// TIA Portal project "FABRICA DE TAPAS - TRANSPORTE -TUNEL DE ENFRIAMIENTO" (V17) (continued)
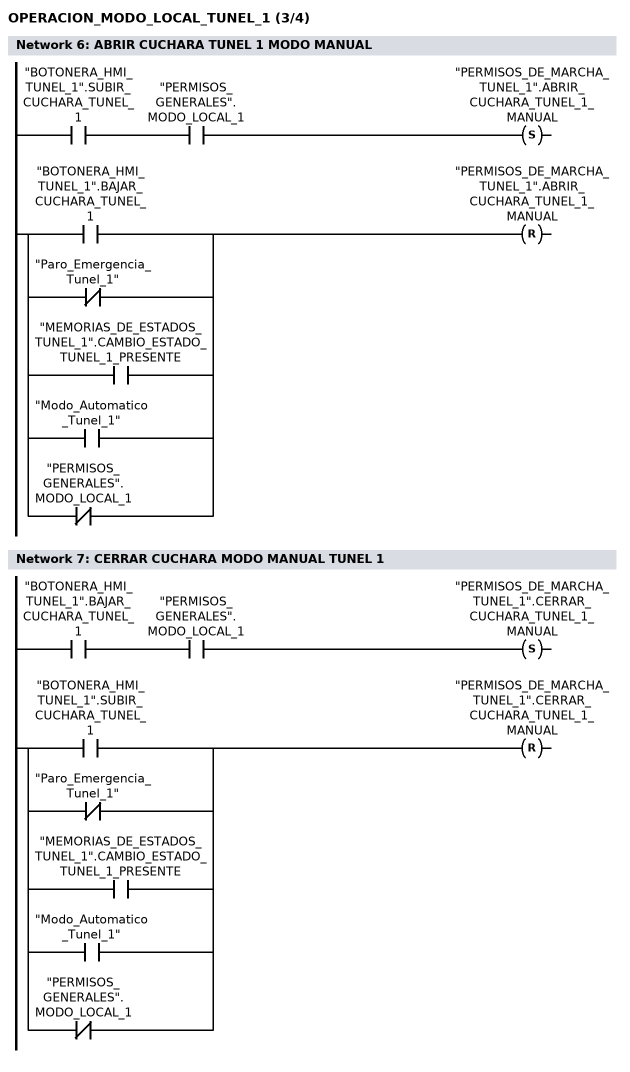
   RUNG wire#powerrail
      Contact( "BOTONERA_HMI_TUNEL_1".SUBIR_CUCHARA_TUNEL_1 )
      Contact( "PERMISOS_GENERALES".MODO_LOCAL_1 )
      S_Coil( "PERMISOS_DE_MARCHA_TUNEL_1".ABRIR_CUCHARA_TUNEL_1_MANUAL )
   END_RUNG
   RUNG wire#powerrail
      Contact( "BOTONERA_HMI_TUNEL_1".BAJAR_CUCHARA_TUNEL_1 )
      wire#w1
      R_Coil( "PERMISOS_DE_MARCHA_TUNEL_1".ABRIR_CUCHARA_TUNEL_1_MANUAL )
   END_RUNG
   RUNG wire#powerrail
      I_Contact( "Paro_Emergencia_Tunel_1" )
   END_RUNG wire#w1
   RUNG wire#powerrail
      Contact( "MEMORIAS_DE_ESTADOS_TUNEL_1".CAMBIO_ESTADO_TUNEL_1_PRESENTE )
   END_RUNG wire#w1
   RUNG wire#powerrail
      Contact( "Modo_Automatico_Tunel_1" )
   END_RUNG wire#w1
   RUNG wire#powerrail
      I_Contact( "PERMISOS_GENERALES".MODO_LOCAL_1 )
   END_RUNG wire#w1
   // the same network as SCL:
   IF "BOTONERA_HMI_TUNEL_1".SUBIR_CUCHARA_TUNEL_1 AND "PERMISOS_GENERALES".MODO_LOCAL_1 THEN
       "PERMISOS_DE_MARCHA_TUNEL_1".ABRIR_CUCHARA_TUNEL_1_MANUAL := TRUE;
   END_IF;
   IF "BOTONERA_HMI_TUNEL_1".BAJAR_CUCHARA_TUNEL_1 OR NOT "Paro_Emergencia_Tunel_1" OR "MEMORIAS_DE_ESTADOS_TUNEL_1".CAMBIO_ESTADO_TUNEL_1_PRESENTE OR "Modo_Automatico_Tunel_1" OR NOT "PERMISOS_GENERALES".MODO_LOCAL_1 THEN
       "PERMISOS_DE_MARCHA_TUNEL_1".ABRIR_CUCHARA_TUNEL_1_MANUAL := FALSE;
   END_IF;
END_REGION

REGION Network 7: CERRAR CUCHARA MODO MANUAL TUNEL 1
   RUNG wire#powerrail
      Contact( "BOTONERA_HMI_TUNEL_1".BAJAR_CUCHARA_TUNEL_1 )
      Contact( "PERMISOS_GENERALES".MODO_LOCAL_1 )
      S_Coil( "PERMISOS_DE_MARCHA_TUNEL_1".CERRAR_CUCHARA_TUNEL_1_MANUAL )
   END_RUNG
   RUNG wire#powerrail
      Contact( "BOTONERA_HMI_TUNEL_1".SUBIR_CUCHARA_TUNEL_1 )
      wire#w1
      R_Coil( "PERMISOS_DE_MARCHA_TUNEL_1".CERRAR_CUCHARA_TUNEL_1_MANUAL )
   END_RUNG
   RUNG wire#powerrail
      I_Contact( "Paro_Emergencia_Tunel_1" )
   END_RUNG wire#w1
   RUNG wire#powerrail
      Contact( "MEMORIAS_DE_ESTADOS_TUNEL_1".CAMBIO_ESTADO_TUNEL_1_PRESENTE )
   END_RUNG wire#w1
   RUNG wire#powerrail
      Contact( "Modo_Automatico_Tunel_1" )
   END_RUNG wire#w1
   RUNG wire#powerrail
      I_Contact( "PERMISOS_GENERALES".MODO_LOCAL_1 )
   END_RUNG wire#w1
   // the same network as SCL:
   IF "BOTONERA_HMI_TUNEL_1".BAJAR_CUCHARA_TUNEL_1 AND "PERMISOS_GENERALES".MODO_LOCAL_1 THEN
       "PERMISOS_DE_MARCHA_TUNEL_1".CERRAR_CUCHARA_TUNEL_1_MANUAL := TRUE;
   END_IF;
   IF "BOTONERA_HMI_TUNEL_1".SUBIR_CUCHARA_TUNEL_1 OR NOT "Paro_Emergencia_Tunel_1" OR "MEMORIAS_DE_ESTADOS_TUNEL_1".CAMBIO_ESTADO_TUNEL_1_PRESENTE OR "Modo_Automatico_Tunel_1" OR NOT "PERMISOS_GENERALES".MODO_LOCAL_1 THEN
       "PERMISOS_DE_MARCHA_TUNEL_1".CERRAR_CUCHARA_TUNEL_1_MANUAL := FALSE;
   END_IF;
END_REGION

REGION Network 8: MOVER SEPARADOR CAJAS A LA DERECHA DE MODO MANUAL TUNEL 1
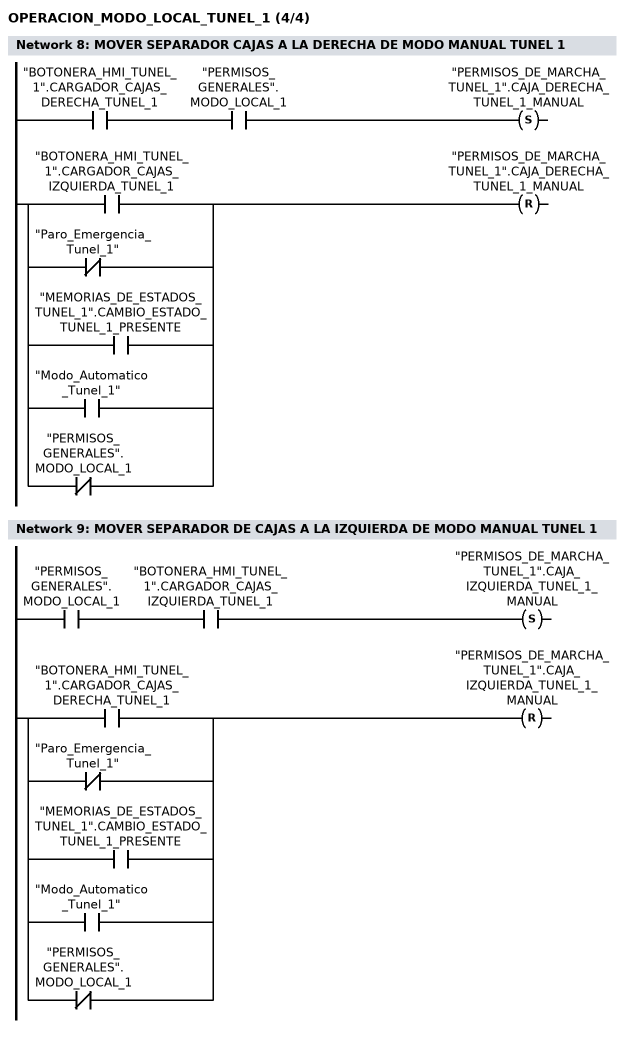
   RUNG wire#powerrail
      Contact( "BOTONERA_HMI_TUNEL_1".CARGADOR_CAJAS_DERECHA_TUNEL_1 )
      Contact( "PERMISOS_GENERALES".MODO_LOCAL_1 )
      S_Coil( "PERMISOS_DE_MARCHA_TUNEL_1".CAJA_DERECHA_TUNEL_1_MANUAL )
   END_RUNG
   RUNG wire#powerrail
      Contact( "BOTONERA_HMI_TUNEL_1".CARGADOR_CAJAS_IZQUIERDA_TUNEL_1 )
      wire#w1
      R_Coil( "PERMISOS_DE_MARCHA_TUNEL_1".CAJA_DERECHA_TUNEL_1_MANUAL )
   END_RUNG
   RUNG wire#powerrail
      I_Contact( "Paro_Emergencia_Tunel_1" )
   END_RUNG wire#w1
   RUNG wire#powerrail
      Contact( "MEMORIAS_DE_ESTADOS_TUNEL_1".CAMBIO_ESTADO_TUNEL_1_PRESENTE )
   END_RUNG wire#w1
   RUNG wire#powerrail
      Contact( "Modo_Automatico_Tunel_1" )
   END_RUNG wire#w1
   RUNG wire#powerrail
      I_Contact( "PERMISOS_GENERALES".MODO_LOCAL_1 )
   END_RUNG wire#w1
   // the same network as SCL:
   IF "BOTONERA_HMI_TUNEL_1".CARGADOR_CAJAS_DERECHA_TUNEL_1 AND "PERMISOS_GENERALES".MODO_LOCAL_1 THEN
       "PERMISOS_DE_MARCHA_TUNEL_1".CAJA_DERECHA_TUNEL_1_MANUAL := TRUE;
   END_IF;
   IF "BOTONERA_HMI_TUNEL_1".CARGADOR_CAJAS_IZQUIERDA_TUNEL_1 OR NOT "Paro_Emergencia_Tunel_1" OR "MEMORIAS_DE_ESTADOS_TUNEL_1".CAMBIO_ESTADO_TUNEL_1_PRESENTE OR "Modo_Automatico_Tunel_1" OR NOT "PERMISOS_GENERALES".MODO_LOCAL_1 THEN
       "PERMISOS_DE_MARCHA_TUNEL_1".CAJA_DERECHA_TUNEL_1_MANUAL := FALSE;
   END_IF;
END_REGION

REGION Network 9: MOVER SEPARADOR DE CAJAS A LA IZQUIERDA DE MODO MANUAL TUNEL 1
   RUNG wire#powerrail
      Contact( "PERMISOS_GENERALES".MODO_LOCAL_1 )
      Contact( "BOTONERA_HMI_TUNEL_1".CARGADOR_CAJAS_IZQUIERDA_TUNEL_1 )
      S_Coil( "PERMISOS_DE_MARCHA_TUNEL_1".CAJA_IZQUIERDA_TUNEL_1_MANUAL )
   END_RUNG
   RUNG wire#powerrail
      Contact( "BOTONERA_HMI_TUNEL_1".CARGADOR_CAJAS_DERECHA_TUNEL_1 )
      wire#w1
      R_Coil( "PERMISOS_DE_MARCHA_TUNEL_1".CAJA_IZQUIERDA_TUNEL_1_MANUAL )
   END_RUNG
   RUNG wire#powerrail
      I_Contact( "Paro_Emergencia_Tunel_1" )
   END_RUNG wire#w1
   RUNG wire#powerrail
      Contact( "MEMORIAS_DE_ESTADOS_TUNEL_1".CAMBIO_ESTADO_TUNEL_1_PRESENTE )
   END_RUNG wire#w1
   RUNG wire#powerrail
      Contact( "Modo_Automatico_Tunel_1" )
   END_RUNG wire#w1
   RUNG wire#powerrail
      I_Contact( "PERMISOS_GENERALES".MODO_LOCAL_1 )
   END_RUNG wire#w1
   // the same network as SCL:
   IF "PERMISOS_GENERALES".MODO_LOCAL_1 AND "BOTONERA_HMI_TUNEL_1".CARGADOR_CAJAS_IZQUIERDA_TUNEL_1 THEN
       "PERMISOS_DE_MARCHA_TUNEL_1".CAJA_IZQUIERDA_TUNEL_1_MANUAL := TRUE;
   END_IF;
   IF "BOTONERA_HMI_TUNEL_1".CARGADOR_CAJAS_DERECHA_TUNEL_1 OR NOT "Paro_Emergencia_Tunel_1" OR "MEMORIAS_DE_ESTADOS_TUNEL_1".CAMBIO_ESTADO_TUNEL_1_PRESENTE OR "Modo_Automatico_Tunel_1" OR NOT "PERMISOS_GENERALES".MODO_LOCAL_1 THEN
       "PERMISOS_DE_MARCHA_TUNEL_1".CAJA_IZQUIERDA_TUNEL_1_MANUAL := FALSE;
   END_IF;
END_REGION
END_FUNCTION

FUNCTION "OPERACION_MODO_LOCAL_TUNEL_2" : Void   // FC4, LAD
{ S7_Optimized_Access := 'TRUE' }
VERSION : 0.1
BEGIN

REGION Network 1
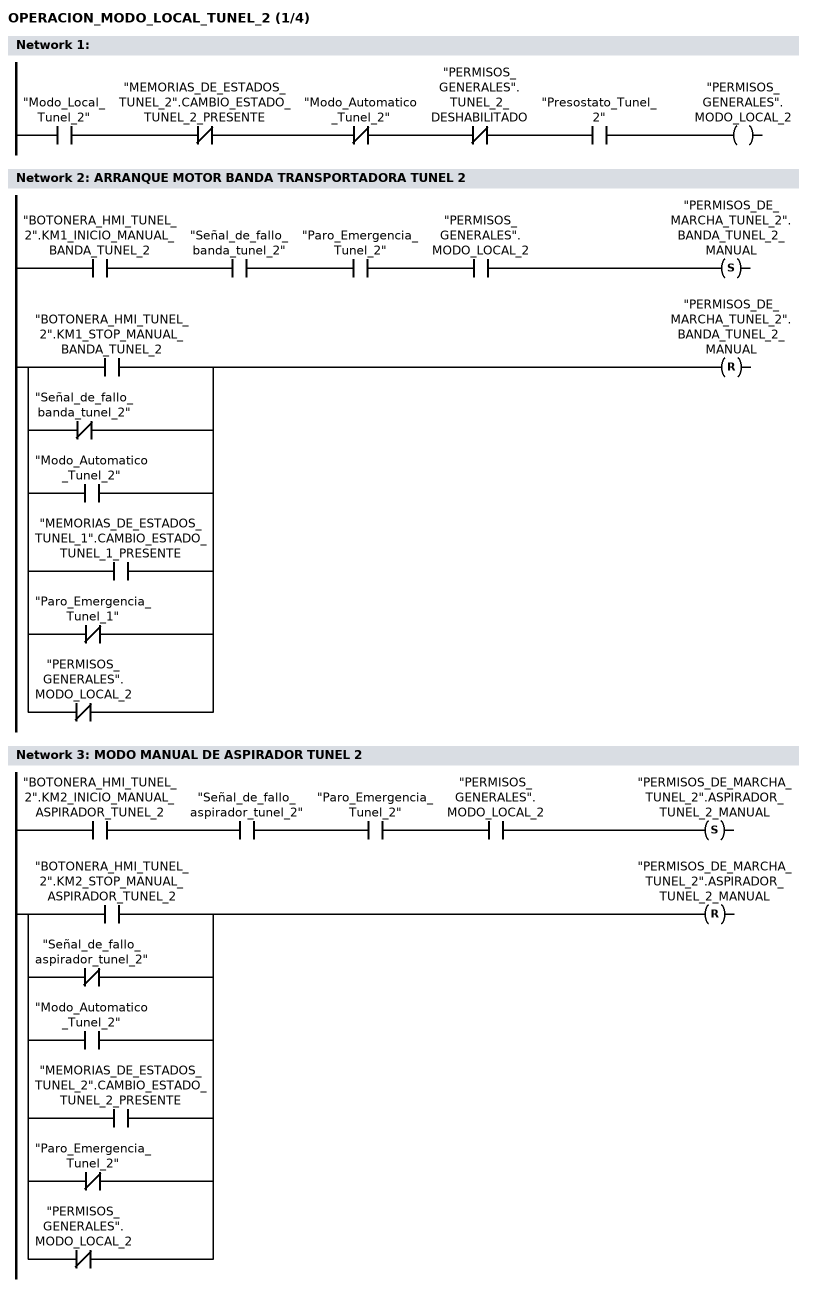
   RUNG wire#powerrail
      Contact( "Modo_Local_Tunel_2" )
      I_Contact( "MEMORIAS_DE_ESTADOS_TUNEL_2".CAMBIO_ESTADO_TUNEL_2_PRESENTE )
      I_Contact( "Modo_Automatico_Tunel_2" )
      I_Contact( "PERMISOS_GENERALES".TUNEL_2_DESHABILITADO )
      Contact( "Presostato_Tunel_2" )
      Coil( "PERMISOS_GENERALES".MODO_LOCAL_2 )
   END_RUNG
   // the same network as SCL:
   "PERMISOS_GENERALES".MODO_LOCAL_2 := "Modo_Local_Tunel_2" AND NOT "MEMORIAS_DE_ESTADOS_TUNEL_2".CAMBIO_ESTADO_TUNEL_2_PRESENTE AND NOT "Modo_Automatico_Tunel_2" AND NOT "PERMISOS_GENERALES".TUNEL_2_DESHABILITADO AND "Presostato_Tunel_2";
END_REGION

REGION Network 2: ARRANQUE MOTOR BANDA TRANSPORTADORA TUNEL 2
   RUNG wire#powerrail
      Contact( "BOTONERA_HMI_TUNEL_2".KM1_INICIO_MANUAL_BANDA_TUNEL_2 )
      Contact( "Señal_de_fallo_banda_tunel_2" )
      Contact( "Paro_Emergencia_Tunel_2" )
      Contact( "PERMISOS_GENERALES".MODO_LOCAL_2 )
      S_Coil( "PERMISOS_DE_MARCHA_TUNEL_2".BANDA_TUNEL_2_MANUAL )
   END_RUNG
   RUNG wire#powerrail
      Contact( "BOTONERA_HMI_TUNEL_2".KM1_STOP_MANUAL_BANDA_TUNEL_2 )
      wire#w1
      R_Coil( "PERMISOS_DE_MARCHA_TUNEL_2".BANDA_TUNEL_2_MANUAL )
   END_RUNG
   RUNG wire#powerrail
      I_Contact( "Señal_de_fallo_banda_tunel_2" )
   END_RUNG wire#w1
   RUNG wire#powerrail
      Contact( "Modo_Automatico_Tunel_2" )
   END_RUNG wire#w1
   RUNG wire#powerrail
      Contact( "MEMORIAS_DE_ESTADOS_TUNEL_1".CAMBIO_ESTADO_TUNEL_1_PRESENTE )
   END_RUNG wire#w1
   RUNG wire#powerrail
      I_Contact( "Paro_Emergencia_Tunel_1" )
   END_RUNG wire#w1
   RUNG wire#powerrail
      I_Contact( "PERMISOS_GENERALES".MODO_LOCAL_2 )
   END_RUNG wire#w1
   // the same network as SCL:
   IF "BOTONERA_HMI_TUNEL_2".KM1_INICIO_MANUAL_BANDA_TUNEL_2 AND "Señal_de_fallo_banda_tunel_2" AND "Paro_Emergencia_Tunel_2" AND "PERMISOS_GENERALES".MODO_LOCAL_2 THEN
       "PERMISOS_DE_MARCHA_TUNEL_2".BANDA_TUNEL_2_MANUAL := TRUE;
   END_IF;
   IF "BOTONERA_HMI_TUNEL_2".KM1_STOP_MANUAL_BANDA_TUNEL_2 OR NOT "Señal_de_fallo_banda_tunel_2" OR "Modo_Automatico_Tunel_2" OR "MEMORIAS_DE_ESTADOS_TUNEL_1".CAMBIO_ESTADO_TUNEL_1_PRESENTE OR NOT "Paro_Emergencia_Tunel_1" OR NOT "PERMISOS_GENERALES".MODO_LOCAL_2 THEN
       "PERMISOS_DE_MARCHA_TUNEL_2".BANDA_TUNEL_2_MANUAL := FALSE;
   END_IF;
END_REGION

REGION Network 3: MODO MANUAL DE ASPIRADOR TUNEL 2
   RUNG wire#powerrail
      Contact( "BOTONERA_HMI_TUNEL_2".KM2_INICIO_MANUAL_ASPIRADOR_TUNEL_2 )
      Contact( "Señal_de_fallo_aspirador_tunel_2" )
      Contact( "Paro_Emergencia_Tunel_2" )
      Contact( "PERMISOS_GENERALES".MODO_LOCAL_2 )
      S_Coil( "PERMISOS_DE_MARCHA_TUNEL_2".ASPIRADOR_TUNEL_2_MANUAL )
   END_RUNG
   RUNG wire#powerrail
      Contact( "BOTONERA_HMI_TUNEL_2".KM2_STOP_MANUAL_ASPIRADOR_TUNEL_2 )
      wire#w1
      R_Coil( "PERMISOS_DE_MARCHA_TUNEL_2".ASPIRADOR_TUNEL_2_MANUAL )
   END_RUNG
   RUNG wire#powerrail
      I_Contact( "Señal_de_fallo_aspirador_tunel_2" )
   END_RUNG wire#w1
   RUNG wire#powerrail
      Contact( "Modo_Automatico_Tunel_2" )
   END_RUNG wire#w1
   RUNG wire#powerrail
      Contact( "MEMORIAS_DE_ESTADOS_TUNEL_2".CAMBIO_ESTADO_TUNEL_2_PRESENTE )
   END_RUNG wire#w1
   RUNG wire#powerrail
      I_Contact( "Paro_Emergencia_Tunel_2" )
   END_RUNG wire#w1
   RUNG wire#powerrail
      I_Contact( "PERMISOS_GENERALES".MODO_LOCAL_2 )
   END_RUNG wire#w1
   // the same network as SCL:
   IF "BOTONERA_HMI_TUNEL_2".KM2_INICIO_MANUAL_ASPIRADOR_TUNEL_2 AND "Señal_de_fallo_aspirador_tunel_2" AND "Paro_Emergencia_Tunel_2" AND "PERMISOS_GENERALES".MODO_LOCAL_2 THEN
       "PERMISOS_DE_MARCHA_TUNEL_2".ASPIRADOR_TUNEL_2_MANUAL := TRUE;
   END_IF;
   IF "BOTONERA_HMI_TUNEL_2".KM2_STOP_MANUAL_ASPIRADOR_TUNEL_2 OR NOT "Señal_de_fallo_aspirador_tunel_2" OR "Modo_Automatico_Tunel_2" OR "MEMORIAS_DE_ESTADOS_TUNEL_2".CAMBIO_ESTADO_TUNEL_2_PRESENTE OR NOT "Paro_Emergencia_Tunel_2" OR NOT "PERMISOS_GENERALES".MODO_LOCAL_2 THEN
       "PERMISOS_DE_MARCHA_TUNEL_2".ASPIRADOR_TUNEL_2_MANUAL := FALSE;
   END_IF;
END_REGION

REGION Network 4: MODO MANUAL VENTILADOR TUNEL 2
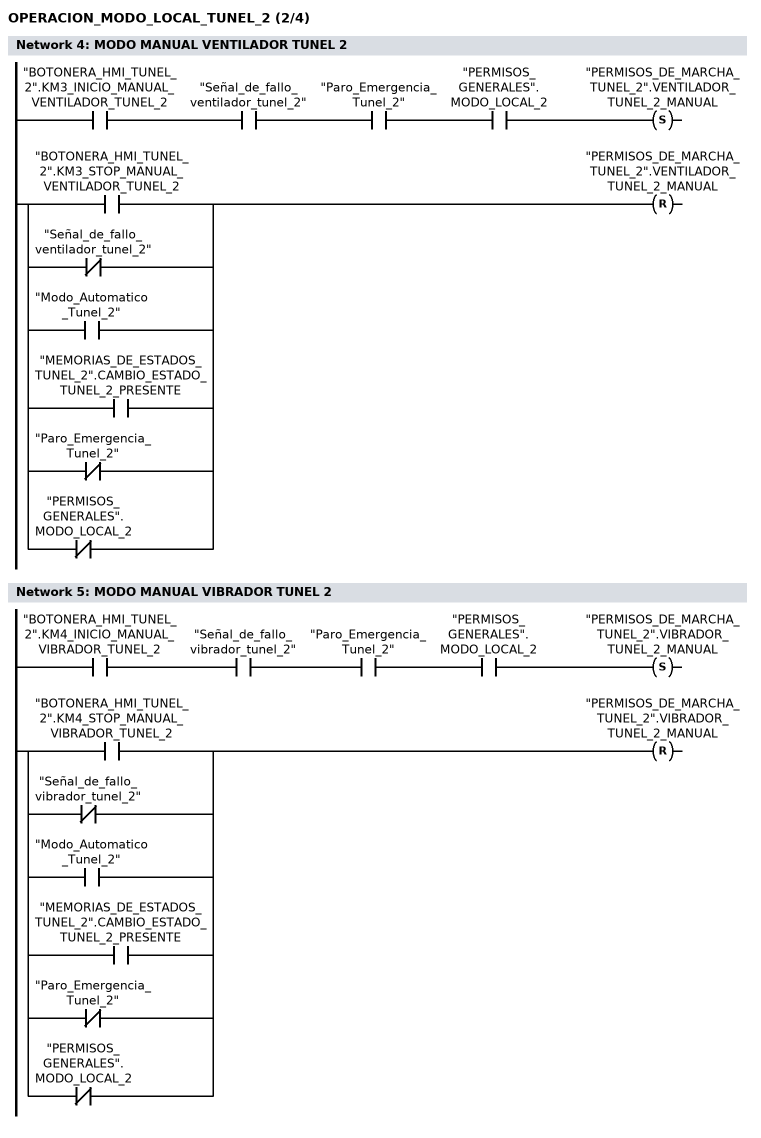
   RUNG wire#powerrail
      Contact( "BOTONERA_HMI_TUNEL_2".KM3_INICIO_MANUAL_VENTILADOR_TUNEL_2 )
      Contact( "Señal_de_fallo_ventilador_tunel_2" )
      Contact( "Paro_Emergencia_Tunel_2" )
      Contact( "PERMISOS_GENERALES".MODO_LOCAL_2 )
      S_Coil( "PERMISOS_DE_MARCHA_TUNEL_2".VENTILADOR_TUNEL_2_MANUAL )
   END_RUNG
   RUNG wire#powerrail
      Contact( "BOTONERA_HMI_TUNEL_2".KM3_STOP_MANUAL_VENTILADOR_TUNEL_2 )
      wire#w1
      R_Coil( "PERMISOS_DE_MARCHA_TUNEL_2".VENTILADOR_TUNEL_2_MANUAL )
   END_RUNG
   RUNG wire#powerrail
      I_Contact( "Señal_de_fallo_ventilador_tunel_2" )
   END_RUNG wire#w1
   RUNG wire#powerrail
      Contact( "Modo_Automatico_Tunel_2" )
   END_RUNG wire#w1
   RUNG wire#powerrail
      Contact( "MEMORIAS_DE_ESTADOS_TUNEL_2".CAMBIO_ESTADO_TUNEL_2_PRESENTE )
   END_RUNG wire#w1
   RUNG wire#powerrail
      I_Contact( "Paro_Emergencia_Tunel_2" )
   END_RUNG wire#w1
   RUNG wire#powerrail
      I_Contact( "PERMISOS_GENERALES".MODO_LOCAL_2 )
   END_RUNG wire#w1
   // the same network as SCL:
   IF "BOTONERA_HMI_TUNEL_2".KM3_INICIO_MANUAL_VENTILADOR_TUNEL_2 AND "Señal_de_fallo_ventilador_tunel_2" AND "Paro_Emergencia_Tunel_2" AND "PERMISOS_GENERALES".MODO_LOCAL_2 THEN
       "PERMISOS_DE_MARCHA_TUNEL_2".VENTILADOR_TUNEL_2_MANUAL := TRUE;
   END_IF;
   IF "BOTONERA_HMI_TUNEL_2".KM3_STOP_MANUAL_VENTILADOR_TUNEL_2 OR NOT "Señal_de_fallo_ventilador_tunel_2" OR "Modo_Automatico_Tunel_2" OR "MEMORIAS_DE_ESTADOS_TUNEL_2".CAMBIO_ESTADO_TUNEL_2_PRESENTE OR NOT "Paro_Emergencia_Tunel_2" OR NOT "PERMISOS_GENERALES".MODO_LOCAL_2 THEN
       "PERMISOS_DE_MARCHA_TUNEL_2".VENTILADOR_TUNEL_2_MANUAL := FALSE;
   END_IF;
END_REGION

REGION Network 5: MODO MANUAL VIBRADOR TUNEL 2
   RUNG wire#powerrail
      Contact( "BOTONERA_HMI_TUNEL_2".KM4_INICIO_MANUAL_VIBRADOR_TUNEL_2 )
      Contact( "Señal_de_fallo_vibrador_tunel_2" )
      Contact( "Paro_Emergencia_Tunel_2" )
      Contact( "PERMISOS_GENERALES".MODO_LOCAL_2 )
      S_Coil( "PERMISOS_DE_MARCHA_TUNEL_2".VIBRADOR_TUNEL_2_MANUAL )
   END_RUNG
   RUNG wire#powerrail
      Contact( "BOTONERA_HMI_TUNEL_2".KM4_STOP_MANUAL_VIBRADOR_TUNEL_2 )
      wire#w1
      R_Coil( "PERMISOS_DE_MARCHA_TUNEL_2".VIBRADOR_TUNEL_2_MANUAL )
   END_RUNG
   RUNG wire#powerrail
      I_Contact( "Señal_de_fallo_vibrador_tunel_2" )
   END_RUNG wire#w1
   RUNG wire#powerrail
      Contact( "Modo_Automatico_Tunel_2" )
   END_RUNG wire#w1
   RUNG wire#powerrail
      Contact( "MEMORIAS_DE_ESTADOS_TUNEL_2".CAMBIO_ESTADO_TUNEL_2_PRESENTE )
   END_RUNG wire#w1
   RUNG wire#powerrail
      I_Contact( "Paro_Emergencia_Tunel_2" )
   END_RUNG wire#w1
   RUNG wire#powerrail
      I_Contact( "PERMISOS_GENERALES".MODO_LOCAL_2 )
   END_RUNG wire#w1
   // the same network as SCL:
   IF "BOTONERA_HMI_TUNEL_2".KM4_INICIO_MANUAL_VIBRADOR_TUNEL_2 AND "Señal_de_fallo_vibrador_tunel_2" AND "Paro_Emergencia_Tunel_2" AND "PERMISOS_GENERALES".MODO_LOCAL_2 THEN
       "PERMISOS_DE_MARCHA_TUNEL_2".VIBRADOR_TUNEL_2_MANUAL := TRUE;
   END_IF;
   IF "BOTONERA_HMI_TUNEL_2".KM4_STOP_MANUAL_VIBRADOR_TUNEL_2 OR NOT "Señal_de_fallo_vibrador_tunel_2" OR "Modo_Automatico_Tunel_2" OR "MEMORIAS_DE_ESTADOS_TUNEL_2".CAMBIO_ESTADO_TUNEL_2_PRESENTE OR NOT "Paro_Emergencia_Tunel_2" OR NOT "PERMISOS_GENERALES".MODO_LOCAL_2 THEN
       "PERMISOS_DE_MARCHA_TUNEL_2".VIBRADOR_TUNEL_2_MANUAL := FALSE;
   END_IF;
END_REGION

REGION Network 6: ABRIR CUCHARA TUNEL 2 MODO MANUAL
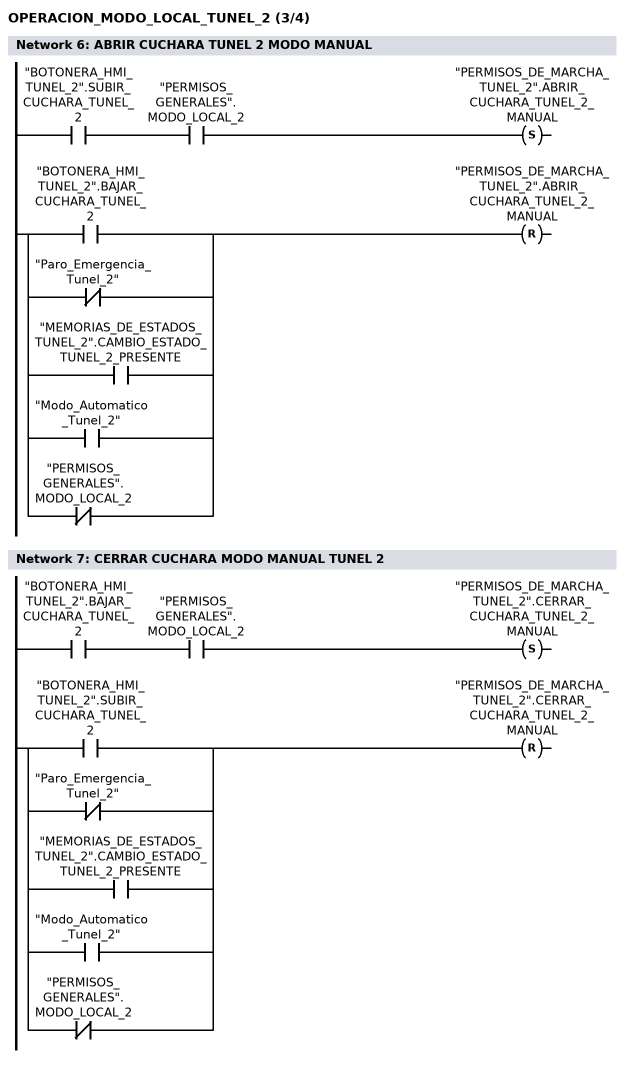
   RUNG wire#powerrail
      Contact( "BOTONERA_HMI_TUNEL_2".SUBIR_CUCHARA_TUNEL_2 )
      Contact( "PERMISOS_GENERALES".MODO_LOCAL_2 )
      S_Coil( "PERMISOS_DE_MARCHA_TUNEL_2".ABRIR_CUCHARA_TUNEL_2_MANUAL )
   END_RUNG
   RUNG wire#powerrail
      Contact( "BOTONERA_HMI_TUNEL_2".BAJAR_CUCHARA_TUNEL_2 )
      wire#w1
      R_Coil( "PERMISOS_DE_MARCHA_TUNEL_2".ABRIR_CUCHARA_TUNEL_2_MANUAL )
   END_RUNG
   RUNG wire#powerrail
      I_Contact( "Paro_Emergencia_Tunel_2" )
   END_RUNG wire#w1
   RUNG wire#powerrail
      Contact( "MEMORIAS_DE_ESTADOS_TUNEL_2".CAMBIO_ESTADO_TUNEL_2_PRESENTE )
   END_RUNG wire#w1
   RUNG wire#powerrail
      Contact( "Modo_Automatico_Tunel_2" )
   END_RUNG wire#w1
   RUNG wire#powerrail
      I_Contact( "PERMISOS_GENERALES".MODO_LOCAL_2 )
   END_RUNG wire#w1
   // the same network as SCL:
   IF "BOTONERA_HMI_TUNEL_2".SUBIR_CUCHARA_TUNEL_2 AND "PERMISOS_GENERALES".MODO_LOCAL_2 THEN
       "PERMISOS_DE_MARCHA_TUNEL_2".ABRIR_CUCHARA_TUNEL_2_MANUAL := TRUE;
   END_IF;
   IF "BOTONERA_HMI_TUNEL_2".BAJAR_CUCHARA_TUNEL_2 OR NOT "Paro_Emergencia_Tunel_2" OR "MEMORIAS_DE_ESTADOS_TUNEL_2".CAMBIO_ESTADO_TUNEL_2_PRESENTE OR "Modo_Automatico_Tunel_2" OR NOT "PERMISOS_GENERALES".MODO_LOCAL_2 THEN
       "PERMISOS_DE_MARCHA_TUNEL_2".ABRIR_CUCHARA_TUNEL_2_MANUAL := FALSE;
   END_IF;
END_REGION

REGION Network 7: CERRAR CUCHARA MODO MANUAL TUNEL 2
   RUNG wire#powerrail
      Contact( "BOTONERA_HMI_TUNEL_2".BAJAR_CUCHARA_TUNEL_2 )
      Contact( "PERMISOS_GENERALES".MODO_LOCAL_2 )
      S_Coil( "PERMISOS_DE_MARCHA_TUNEL_2".CERRAR_CUCHARA_TUNEL_2_MANUAL )
   END_RUNG
   RUNG wire#powerrail
      Contact( "BOTONERA_HMI_TUNEL_2".SUBIR_CUCHARA_TUNEL_2 )
      wire#w1
      R_Coil( "PERMISOS_DE_MARCHA_TUNEL_2".CERRAR_CUCHARA_TUNEL_2_MANUAL )
   END_RUNG
   RUNG wire#powerrail
      I_Contact( "Paro_Emergencia_Tunel_2" )
   END_RUNG wire#w1
   RUNG wire#powerrail
      Contact( "MEMORIAS_DE_ESTADOS_TUNEL_2".CAMBIO_ESTADO_TUNEL_2_PRESENTE )
   END_RUNG wire#w1
   RUNG wire#powerrail
      Contact( "Modo_Automatico_Tunel_2" )
   END_RUNG wire#w1
   RUNG wire#powerrail
      I_Contact( "PERMISOS_GENERALES".MODO_LOCAL_2 )
   END_RUNG wire#w1
   // the same network as SCL:
   IF "BOTONERA_HMI_TUNEL_2".BAJAR_CUCHARA_TUNEL_2 AND "PERMISOS_GENERALES".MODO_LOCAL_2 THEN
       "PERMISOS_DE_MARCHA_TUNEL_2".CERRAR_CUCHARA_TUNEL_2_MANUAL := TRUE;
   END_IF;
   IF "BOTONERA_HMI_TUNEL_2".SUBIR_CUCHARA_TUNEL_2 OR NOT "Paro_Emergencia_Tunel_2" OR "MEMORIAS_DE_ESTADOS_TUNEL_2".CAMBIO_ESTADO_TUNEL_2_PRESENTE OR "Modo_Automatico_Tunel_2" OR NOT "PERMISOS_GENERALES".MODO_LOCAL_2 THEN
       "PERMISOS_DE_MARCHA_TUNEL_2".CERRAR_CUCHARA_TUNEL_2_MANUAL := FALSE;
   END_IF;
END_REGION

REGION Network 8: MOVER SEPARADOR CAJAS A LA DERECHA DE MODO MANUAL TUNEL 2
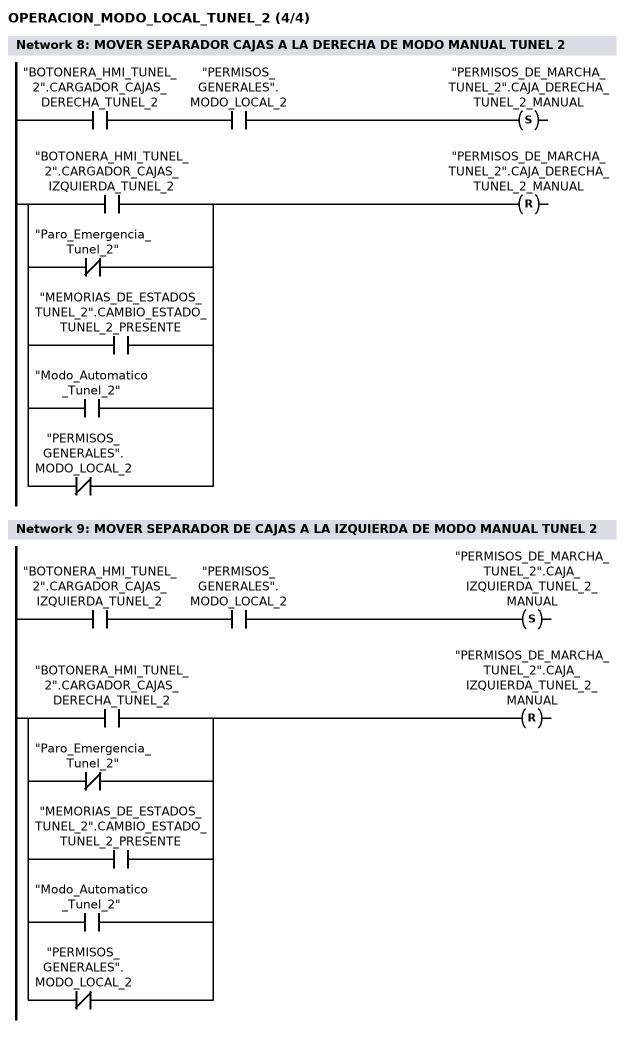
   RUNG wire#powerrail
      Contact( "BOTONERA_HMI_TUNEL_2".CARGADOR_CAJAS_DERECHA_TUNEL_2 )
      Contact( "PERMISOS_GENERALES".MODO_LOCAL_2 )
      S_Coil( "PERMISOS_DE_MARCHA_TUNEL_2".CAJA_DERECHA_TUNEL_2_MANUAL )
   END_RUNG
   RUNG wire#powerrail
      Contact( "BOTONERA_HMI_TUNEL_2".CARGADOR_CAJAS_IZQUIERDA_TUNEL_2 )
      wire#w1
      R_Coil( "PERMISOS_DE_MARCHA_TUNEL_2".CAJA_DERECHA_TUNEL_2_MANUAL )
   END_RUNG
   RUNG wire#powerrail
      I_Contact( "Paro_Emergencia_Tunel_2" )
   END_RUNG wire#w1
   RUNG wire#powerrail
      Contact( "MEMORIAS_DE_ESTADOS_TUNEL_2".CAMBIO_ESTADO_TUNEL_2_PRESENTE )
   END_RUNG wire#w1
   RUNG wire#powerrail
      Contact( "Modo_Automatico_Tunel_2" )
   END_RUNG wire#w1
   RUNG wire#powerrail
      I_Contact( "PERMISOS_GENERALES".MODO_LOCAL_2 )
   END_RUNG wire#w1
   // the same network as SCL:
   IF "BOTONERA_HMI_TUNEL_2".CARGADOR_CAJAS_DERECHA_TUNEL_2 AND "PERMISOS_GENERALES".MODO_LOCAL_2 THEN
       "PERMISOS_DE_MARCHA_TUNEL_2".CAJA_DERECHA_TUNEL_2_MANUAL := TRUE;
   END_IF;
   IF "BOTONERA_HMI_TUNEL_2".CARGADOR_CAJAS_IZQUIERDA_TUNEL_2 OR NOT "Paro_Emergencia_Tunel_2" OR "MEMORIAS_DE_ESTADOS_TUNEL_2".CAMBIO_ESTADO_TUNEL_2_PRESENTE OR "Modo_Automatico_Tunel_2" OR NOT "PERMISOS_GENERALES".MODO_LOCAL_2 THEN
       "PERMISOS_DE_MARCHA_TUNEL_2".CAJA_DERECHA_TUNEL_2_MANUAL := FALSE;
   END_IF;
END_REGION

REGION Network 9: MOVER SEPARADOR DE CAJAS A LA IZQUIERDA DE MODO MANUAL TUNEL 2
   RUNG wire#powerrail
      Contact( "BOTONERA_HMI_TUNEL_2".CARGADOR_CAJAS_IZQUIERDA_TUNEL_2 )
      Contact( "PERMISOS_GENERALES".MODO_LOCAL_2 )
      S_Coil( "PERMISOS_DE_MARCHA_TUNEL_2".CAJA_IZQUIERDA_TUNEL_2_MANUAL )
   END_RUNG
   RUNG wire#powerrail
      Contact( "BOTONERA_HMI_TUNEL_2".CARGADOR_CAJAS_DERECHA_TUNEL_2 )
      wire#w1
      R_Coil( "PERMISOS_DE_MARCHA_TUNEL_2".CAJA_IZQUIERDA_TUNEL_2_MANUAL )
   END_RUNG
   RUNG wire#powerrail
      I_Contact( "Paro_Emergencia_Tunel_2" )
   END_RUNG wire#w1
   RUNG wire#powerrail
      Contact( "MEMORIAS_DE_ESTADOS_TUNEL_2".CAMBIO_ESTADO_TUNEL_2_PRESENTE )
   END_RUNG wire#w1
   RUNG wire#powerrail
      Contact( "Modo_Automatico_Tunel_2" )
   END_RUNG wire#w1
   RUNG wire#powerrail
      I_Contact( "PERMISOS_GENERALES".MODO_LOCAL_2 )
   END_RUNG wire#w1
   // the same network as SCL:
   IF "BOTONERA_HMI_TUNEL_2".CARGADOR_CAJAS_IZQUIERDA_TUNEL_2 AND "PERMISOS_GENERALES".MODO_LOCAL_2 THEN
       "PERMISOS_DE_MARCHA_TUNEL_2".CAJA_IZQUIERDA_TUNEL_2_MANUAL := TRUE;
   END_IF;
   IF "BOTONERA_HMI_TUNEL_2".CARGADOR_CAJAS_DERECHA_TUNEL_2 OR NOT "Paro_Emergencia_Tunel_2" OR "MEMORIAS_DE_ESTADOS_TUNEL_2".CAMBIO_ESTADO_TUNEL_2_PRESENTE OR "Modo_Automatico_Tunel_2" OR NOT "PERMISOS_GENERALES".MODO_LOCAL_2 THEN
       "PERMISOS_DE_MARCHA_TUNEL_2".CAJA_IZQUIERDA_TUNEL_2_MANUAL := FALSE;
   END_IF;
END_REGION
END_FUNCTION

FUNCTION "OPERACION_MANUAL_TRANSPORTE" : Void   // FC5, LAD
{ S7_Optimized_Access := 'TRUE' }
VERSION : 0.1
BEGIN

REGION Network 1
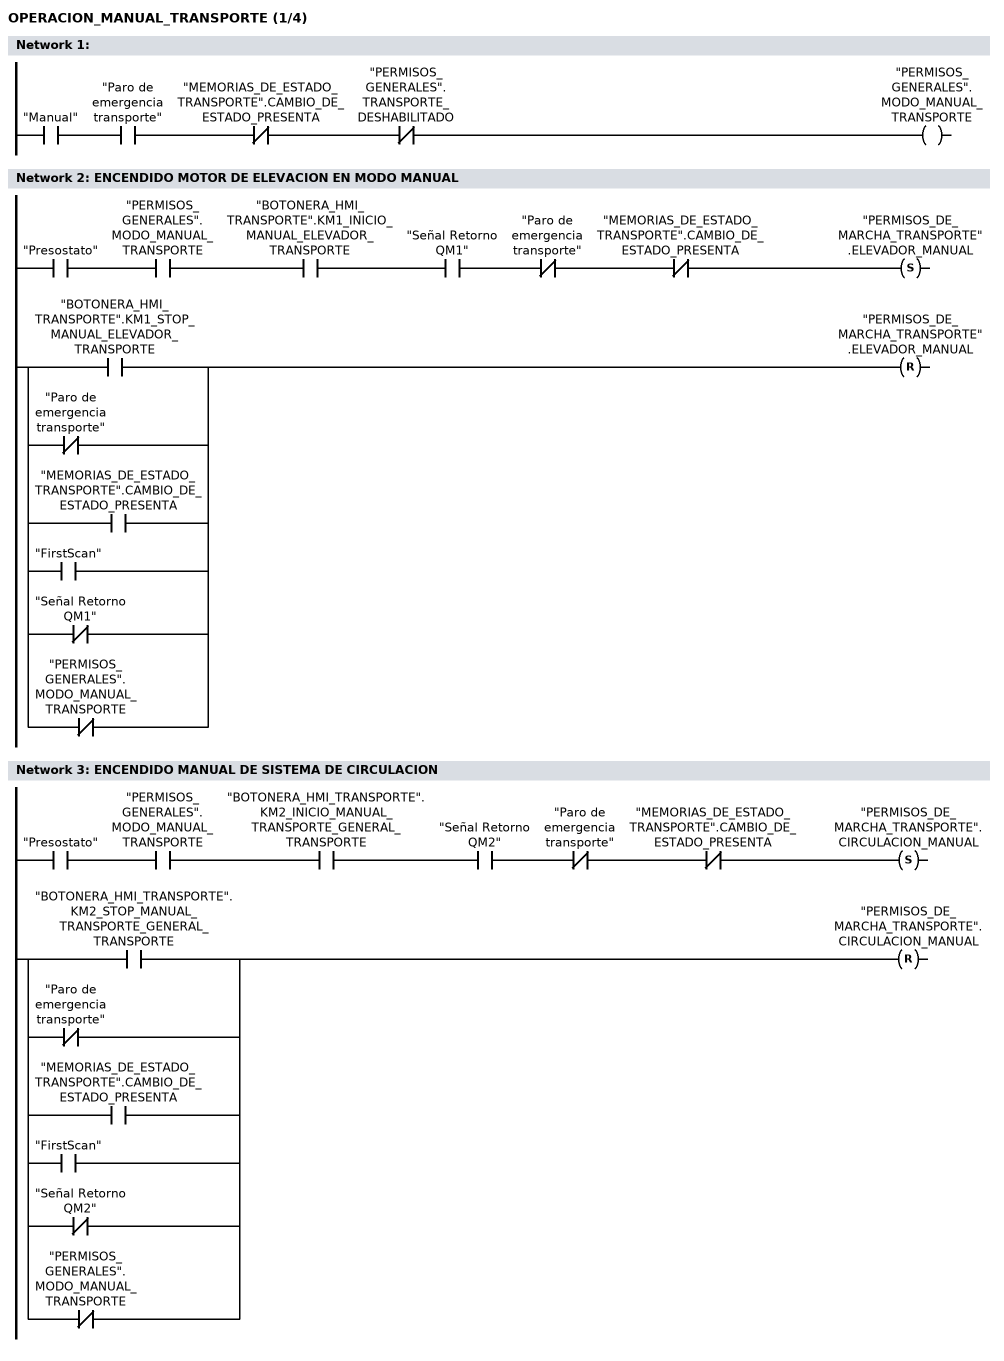
   RUNG wire#powerrail
      Contact( "Manual" )
      Contact( "Paro de emergencia transporte" )
      I_Contact( "MEMORIAS_DE_ESTADO_TRANSPORTE".CAMBIO_DE_ESTADO_PRESENTA )
      I_Contact( "PERMISOS_GENERALES".TRANSPORTE_DESHABILITADO )
      Coil( "PERMISOS_GENERALES".MODO_MANUAL_TRANSPORTE )
   END_RUNG
   // the same network as SCL:
   "PERMISOS_GENERALES".MODO_MANUAL_TRANSPORTE := "Manual" AND "Paro de emergencia transporte" AND NOT "MEMORIAS_DE_ESTADO_TRANSPORTE".CAMBIO_DE_ESTADO_PRESENTA AND NOT "PERMISOS_GENERALES".TRANSPORTE_DESHABILITADO;
END_REGION

REGION Network 2: ENCENDIDO MOTOR DE ELEVACION EN MODO MANUAL
   RUNG wire#powerrail
      Contact( "Presostato" )
      Contact( "PERMISOS_GENERALES".MODO_MANUAL_TRANSPORTE )
      Contact( "BOTONERA_HMI_TRANSPORTE".KM1_INICIO_MANUAL_ELEVADOR_TRANSPORTE )
      Contact( "Señal Retorno QM1" )
      I_Contact( "Paro de emergencia transporte" )
      I_Contact( "MEMORIAS_DE_ESTADO_TRANSPORTE".CAMBIO_DE_ESTADO_PRESENTA )
      S_Coil( "PERMISOS_DE_MARCHA_TRANSPORTE".ELEVADOR_MANUAL )
   END_RUNG
   RUNG wire#powerrail
      Contact( "BOTONERA_HMI_TRANSPORTE".KM1_STOP_MANUAL_ELEVADOR_TRANSPORTE )
      wire#w1
      R_Coil( "PERMISOS_DE_MARCHA_TRANSPORTE".ELEVADOR_MANUAL )
   END_RUNG
   RUNG wire#powerrail
      I_Contact( "Paro de emergencia transporte" )
   END_RUNG wire#w1
   RUNG wire#powerrail
      Contact( "MEMORIAS_DE_ESTADO_TRANSPORTE".CAMBIO_DE_ESTADO_PRESENTA )
   END_RUNG wire#w1
   RUNG wire#powerrail
      Contact( "FirstScan" )
   END_RUNG wire#w1
   RUNG wire#powerrail
      I_Contact( "Señal Retorno QM1" )
   END_RUNG wire#w1
   RUNG wire#powerrail
      I_Contact( "PERMISOS_GENERALES".MODO_MANUAL_TRANSPORTE )
   END_RUNG wire#w1
   // the same network as SCL:
   IF "Presostato" AND "PERMISOS_GENERALES".MODO_MANUAL_TRANSPORTE AND "BOTONERA_HMI_TRANSPORTE".KM1_INICIO_MANUAL_ELEVADOR_TRANSPORTE AND "Señal Retorno QM1" AND NOT "Paro de emergencia transporte" AND NOT "MEMORIAS_DE_ESTADO_TRANSPORTE".CAMBIO_DE_ESTADO_PRESENTA THEN
       "PERMISOS_DE_MARCHA_TRANSPORTE".ELEVADOR_MANUAL := TRUE;
   END_IF;
   IF "BOTONERA_HMI_TRANSPORTE".KM1_STOP_MANUAL_ELEVADOR_TRANSPORTE OR NOT "Paro de emergencia transporte" OR "MEMORIAS_DE_ESTADO_TRANSPORTE".CAMBIO_DE_ESTADO_PRESENTA OR "FirstScan" OR NOT "Señal Retorno QM1" OR NOT "PERMISOS_GENERALES".MODO_MANUAL_TRANSPORTE THEN
       "PERMISOS_DE_MARCHA_TRANSPORTE".ELEVADOR_MANUAL := FALSE;
   END_IF;
END_REGION

REGION Network 3: ENCENDIDO MANUAL DE SISTEMA DE CIRCULACION
   RUNG wire#powerrail
      Contact( "Presostato" )
      Contact( "PERMISOS_GENERALES".MODO_MANUAL_TRANSPORTE )
      Contact( "BOTONERA_HMI_TRANSPORTE".KM2_INICIO_MANUAL_TRANSPORTE_GENERAL_TRANSPORTE )
      Contact( "Señal Retorno QM2" )
      I_Contact( "Paro de emergencia transporte" )
      I_Contact( "MEMORIAS_DE_ESTADO_TRANSPORTE".CAMBIO_DE_ESTADO_PRESENTA )
      S_Coil( "PERMISOS_DE_MARCHA_TRANSPORTE".CIRCULACION_MANUAL )
   END_RUNG
   RUNG wire#powerrail
      Contact( "BOTONERA_HMI_TRANSPORTE".KM2_STOP_MANUAL_TRANSPORTE_GENERAL_TRANSPORTE )
      wire#w1
      R_Coil( "PERMISOS_DE_MARCHA_TRANSPORTE".CIRCULACION_MANUAL )
   END_RUNG
   RUNG wire#powerrail
      I_Contact( "Paro de emergencia transporte" )
   END_RUNG wire#w1
   RUNG wire#powerrail
      Contact( "MEMORIAS_DE_ESTADO_TRANSPORTE".CAMBIO_DE_ESTADO_PRESENTA )
   END_RUNG wire#w1
   RUNG wire#powerrail
      Contact( "FirstScan" )
   END_RUNG wire#w1
   RUNG wire#powerrail
      I_Contact( "Señal Retorno QM2" )
   END_RUNG wire#w1
   RUNG wire#powerrail
      I_Contact( "PERMISOS_GENERALES".MODO_MANUAL_TRANSPORTE )
   END_RUNG wire#w1
   // the same network as SCL:
   IF "Presostato" AND "PERMISOS_GENERALES".MODO_MANUAL_TRANSPORTE AND "BOTONERA_HMI_TRANSPORTE".KM2_INICIO_MANUAL_TRANSPORTE_GENERAL_TRANSPORTE AND "Señal Retorno QM2" AND NOT "Paro de emergencia transporte" AND NOT "MEMORIAS_DE_ESTADO_TRANSPORTE".CAMBIO_DE_ESTADO_PRESENTA THEN
       "PERMISOS_DE_MARCHA_TRANSPORTE".CIRCULACION_MANUAL := TRUE;
   END_IF;
   IF "BOTONERA_HMI_TRANSPORTE".KM2_STOP_MANUAL_TRANSPORTE_GENERAL_TRANSPORTE OR NOT "Paro de emergencia transporte" OR "MEMORIAS_DE_ESTADO_TRANSPORTE".CAMBIO_DE_ESTADO_PRESENTA OR "FirstScan" OR NOT "Señal Retorno QM2" OR NOT "PERMISOS_GENERALES".MODO_MANUAL_TRANSPORTE THEN
       "PERMISOS_DE_MARCHA_TRANSPORTE".CIRCULACION_MANUAL := FALSE;
   END_IF;
END_REGION

REGION Network 4: LLENADO DE TOLVA RESERVA